DATA_BLOCK "DB_CrossCut_3_HMI"   // DB2078
{ S7_Optimized_Access := 'FALSE' }
VERSION : 0.1
   VAR
      tALM : Struct   // HMI Alarms
         tE : Struct   // Emergency alarms
            xLocON : Bool;   // KE.Local emergency ON {X|X|X|X|O}
            xLocal1 : Bool;   // SB.Local emergency push button 1 {X|X|X|X|O}
            xLocal2 : Bool;   // SB.Local emergency push button 2 {X|X|X|X|O}
            xLocal3 : Bool;   // SB.Local emergency push button 3 {X|X|X|X|O}
            xSpare_4 : Bool;
            xSpare_5 : Bool;
            xSpare_6 : Bool;
            xSpare_7 : Bool;
            xSpare_8 : Bool;
            xSpare_9 : Bool;
            xSpare_10 : Bool;
            xSpare_11 : Bool;
            xSpare_12 : Bool;
            xSpare_13 : Bool;
            xSpare_14 : Bool;
            xSpare_15 : Bool;
            xSpare_16 : Bool;
            xSpare_17 : Bool;
            xSpare_18 : Bool;
            xSpare_19 : Bool;
            xSpare_20 : Bool;
            xSpare_21 : Bool;
            xSpare_22 : Bool;
            xSpare_23 : Bool;
            xSpare_24 : Bool;
            xSpare_25 : Bool;
            xSpare_26 : Bool;
            xSpare_27 : Bool;
            xSpare_28 : Bool;
            xSpare_29 : Bool;
            xSpare_30 : Bool;
            xSpare_31 : Bool;
         END_STRUCT;
         tS : Struct   // Stopping faults
            xAxisNotAvail : Bool;   // AZ.Axis not available {X|X|X|X|O}
            xInpInstallation : Bool;   // L+.Input power supply ON {X|X|X|X|O}
            xAuxPower : Bool;   // L+.Auxiliary power supple set-in {X|X|X|X|O}
            xAreaSafety : Bool;   // KE.Area safety {X|X|X|X|O}
            xOverstroke : Bool;   // KA.Carriage overstroke {X|X|X|X|O}
            xExternInputPower : Bool;   // L+.External input power supply {X|X|X|X|O}
            xCarriageCutOut : Bool;   // QM.Carriage translation overload {X|X|X|X|O}
            xDriveTrip : Bool;   // AZ.Drive trip {X|X|X|X|O}
            xDriveNotEnabled : Bool;   // AZ.Drive not enabled {X|X|X|X|O}
            xAxisNotReady : Bool;   // AZ.Axis not ready {X|X|X|X|O}
            xDriveNotReady : Bool;   // AZ.Drive not ready {X|X|X|X|O}
            xAxisNotSyncro : Bool;   // AZ.Axis not syncronized {X|X|X|X|O}
            xSpare_12 : Bool;
            xSpare_13 : Bool;
            xSpare_14 : Bool;
            xSpare_15 : Bool;
            xSpare_16 : Bool;
            xSpare_17 : Bool;
            xSpare_18 : Bool;
            xSpare_19 : Bool;
            xSpare_20 : Bool;
            xSpare_21 : Bool;
            xSpare_22 : Bool;
            xSpare_23 : Bool;
            xSpare_24 : Bool;
            xSpare_25 : Bool;
            xSpare_26 : Bool;
            xSpare_27 : Bool;
            xSpare_28 : Bool;
            xSpare_29 : Bool;
            xSpare_30 : Bool;
            xSpare_31 : Bool;
         END_STRUCT;
         tF : Struct   // Faults
            xSpare_0 : Bool;
            xSpare_1 : Bool;
            xSpare_2 : Bool;
            xSpare_3 : Bool;
            xSpare_4 : Bool;
            xSpare_5 : Bool;
            xSpare_6 : Bool;
            xSpare_7 : Bool;
            xSpare_8 : Bool;
            xSpare_9 : Bool;
            xSpare_10 : Bool;
            xSpare_11 : Bool;
            xSpare_12 : Bool;
            xSpare_13 : Bool;
            xSpare_14 : Bool;
            xSpare_15 : Bool;
            xSpare_16 : Bool;
            xSpare_17 : Bool;
            xSpare_18 : Bool;
            xSpare_19 : Bool;
            xSpare_20 : Bool;
            xSpare_21 : Bool;
            xSpare_22 : Bool;
            xSpare_23 : Bool;
            xSpare_24 : Bool;
            xSpare_25 : Bool;
            xSpare_26 : Bool;
            xSpare_27 : Bool;
            xSpare_28 : Bool;
            xSpare_29 : Bool;
            xSpare_30 : Bool;
            xSpare_31 : Bool;
         END_STRUCT;
         tW : Struct   // Warnings
            xSpare_0 : Bool;
            xSpare_1 : Bool;
            xSpare_2 : Bool;
            xSpare_3 : Bool;
            xSpare_4 : Bool;
            xSpare_5 : Bool;
            xSpare_6 : Bool;
            xSpare_7 : Bool;
            xSpare_8 : Bool;
            xSpare_9 : Bool;
            xSpare_10 : Bool;
            xSpare_11 : Bool;
            xSpare_12 : Bool;
            xSpare_13 : Bool;
            xSpare_14 : Bool;
            xSpare_15 : Bool;
            xSpare_16 : Bool;
            xSpare_17 : Bool;
            xSpare_18 : Bool;
            xSpare_19 : Bool;
            xSpare_20 : Bool;
            xSpare_21 : Bool;
            xSpare_22 : Bool;
            xSpare_23 : Bool;
            xSpare_24 : Bool;
            xSpare_25 : Bool;
            xSpare_26 : Bool;
            xSpare_27 : Bool;
            xSpare_28 : Bool;
            xSpare_29 : Bool;
            xSpare_30 : Bool;
            xSpare_31 : Bool;
         END_STRUCT;
      END_STRUCT;
      tHMR : Struct   // HMI Read
         xSpare0 : Bool;
         xSpare1 : Bool;
         xSpare2 : Bool;
         xSpare3 : Bool;
         xSpare4 : Bool;
         xSpare5 : Bool;
         xSpare6 : Bool;
         xSpare7 : Bool;
         xSpare8 : Bool;
         xSpare9 : Bool;
         xSpare10 : Bool;
         xSpare11 : Bool;
         xSpare12 : Bool;
         xSpare13 : Bool;
         xManualCommandEnabled : Bool;   // Manual Command enabled {x|x|x|x|O}
         xSpare15 : Bool;
         xSpare16 : Bool;
         xSpare17 : Bool;
         xSpare18 : Bool;
         xSpare19 : Bool;
         xSpare20 : Bool;
         xSpare21 : Bool;
         xSpare22 : Bool;
         xSpare23 : Bool;
         xSpare24 : Bool;
         xSpare25 : Bool;
         xSpare26 : Bool;
         xSpare27 : Bool;
         xSpare28 : Bool;
         xSpare29 : Bool;
         xSpare30 : Bool;
         xSpare31 : Bool;
         xSpare : Array[0..15] of Bool;
         iSpare0 : Int;
         iSpare1 : Int;
         iSpare2 : Int;
         iSpare3 : Int;
         iSpare4 : Int;
         iSpare5 : Int;
         iSpare6 : Int;
         iSpare7 : Int;
         iSpare8 : Int;
         iSpare9 : Int;
         iSpare10 : Int;
         iSpare11 : Int;
         iSpare12 : Int;
         iSpare13 : Int;
         iSpare14 : Int;
         iSpare15 : Int;
         iSpare16 : Int;
         dDistanceSnaproll_cmm : DInt;   // Distance from snaproll [mm/100] {mm/100|mm|x|x|M}
         dStatus : DInt;   // XCut actual status (1=Idle 3=Running 7=Faulted) {X|X|X|X|O}
         dXCutActualStatus : DInt;   // XCut actual status (1=Disabled 3=Enabled) {X|X|X|X|O}
         dXCutStatusRequest : DInt;   // XCut status request (1=Disabled 3=Enabled) {X|X|X|X|O}
         dDistanceFromCenterLine_cmm : DInt;   // Distance from center line [mm/100] {mm/100|mm|X|X|O}
         dAngleValue_uDegree : DInt;   // Angle value [°/1000000] {°/1000000|°|X|X|O}
         dActualCutPosRequest : DInt;   // Actual cut position request (1=By operator 2=On gross ribbon 3=On net ribbon 4=On YCut position) {X|X|X|X|O}
         dCarriagePosition_cmm : DInt;   // Actual carriage position [mm/100]
         dSpare8 : DInt;
         dSpare9 : DInt;
         dSpare10 : DInt;
         dSpare11 : DInt;
         dSpare12 : DInt;
         dSpare13 : DInt;
         dSpare14 : DInt;
         dSpare15 : DInt;
         rHeadUsage_km : Real;   // Head usage [Km] {Km|Km|X|X|O}
         rSpare1 : Real;
         rSpare2 : Real;
         rSpare3 : Real;
         rSpare4 : Real;
         rSpare5 : Real;
         rSpare6 : Real;
         rSpare7 : Real;
         rSpare8 : Real;
         tManCmd : Struct
            xManJogFwdFdbk : Bool;   // Manual jog forward feedback {X|X|X|X|O}
            xManJogBckFdbk : Bool;   // Manual jog backward feedback {X|X|X|X|O}
            xManCarriageDownFdbk : Bool;   // Manual carriage down feedback {X|X|X|X|O}
            xManFireONFdbk : Bool;   // Manual fire ON feedback {X|X|X|X|O}
            xManOilONFdbk : Bool;   // Manual oil ON feedback {X|X|X|X|O}
            xSpare5 : Bool;
            xSpare6 : Bool;
            xSpare7 : Bool;
            xSpare8 : Bool;
            xSpare9 : Bool;
            xSpare10 : Bool;
            xSpare11 : Bool;
            xSpare12 : Bool;
            xSpare13 : Bool;
            xSpare14 : Bool;
            xSpare15 : Bool;
            xSpare : Array[0..15] of Bool;
         END_STRUCT;
      END_STRUCT;
      tHMW : Struct   // HMI Write
         xCutBreakEnabled : Bool;   // Cut on glass break enabled {X|X|X|X|O}
         xIncAngleValue : Bool;   // Increment angle value {X|X|X|X|O}
         xDecAngleValue : Bool;   // Decrement angle value {X|X|X|X|O}
         xCalibDistRequest : Bool;   // Calibration distance request {X|X|X|X|O}
         xCalibDiagRequest : Bool;   // Calibration diagonal request {X|X|X|X|O}
         xCutOperator : Bool;   // Cutting position by operator request {X|X|X|X|O}
         xCutGross : Bool;   // Cutting position by gross width position {X|X|X|X|O}
         xCutNet : Bool;   // Cutting position by net width position {X|X|X|X|O}
         xCutYCut : Bool;   // Cutting position by YCut position {X|X|X|X|O}
         xSpare9 : Bool;
         xSpare10 : Bool;
         xSpare11 : Bool;
         xSpare12 : Bool;
         xResetHeadUsage : Bool;   // Reset the head usage {X|X|X|X|O}
         xEnableManualCommand : Bool;   // Enable Disable Manual command {x|x|x|x|O}
         xUpdateDistanceSnaproll : Bool;   // Update distance from snaproll {x|x|x|x|M}
         xUpdateDistCenterLine : Bool;   // Update distance from center line {X|X|X|X|M}
         xUpdateAngleValue : Bool;   // Update angle value {X|X|X|X|M}
         xSpare18 : Bool;
         xSpare19 : Bool;
         xSpare20 : Bool;
         xSpare21 : Bool;
         xSpare22 : Bool;
         xSpare23 : Bool;
         xSpare24 : Bool;
         xSpare25 : Bool;
         xSpare26 : Bool;
         xSpare27 : Bool;
         xSpare28 : Bool;
         xSpare29 : Bool;
         xSpare30 : Bool;
         xSpare31 : Bool;
         xSpare : Array[0..15] of Bool;
         iSpare0 : Int;
         iSpare1 : Int;
         iSpare2 : Int;
         iSpare3 : Int;
         iSpare4 : Int;
         iSpare5 : Int;
         iSpare6 : Int;
         iSpare7 : Int;
         iSpare8 : Int;
         iSpare9 : Int;
         iSpare10 : Int;
         iSpare11 : Int;
         iSpare12 : Int;
         iSpare13 : Int;
         iSpare14 : Int;
         iSpare15 : Int;
         iSpare16 : Int;
         dDistanceSnaproll_cmm : DInt;   // Distance from snaproll [mm/100] {mm/100|mm|1|70000|M}
         dDistanceFromCenterLine_cmm : DInt;   // Distance from center line [mm/100] {mm/100|mm|-3000|0|M}
         dAngleValue_uDegree : DInt;   // Bridge angle value [°/1000000] {°/1000000|°|7|9|M}
         dOperStartCutPos_cmm : DInt;   // Operator start cut position [mm/100] {mm/100|mm|-3000|0|O}
         dOperEndCutPos_cmm : DInt;   // Operator end cut position [mm/100] {mm/100|mm|0|3000|O}
         dDescReactTime_ms : DInt;   // Carriage descent reaction time [ms] {ms|s|0|1|M}
         dRaiseReactTime_ms : DInt;   // Carriage raise reaction time [ms] {ms|s|0|1|M}
         dFireONReactTime_ms : DInt;   // Fire ON reaction time [ms] {ms|s|0|1|M}
         dFireOFFReactTime_ms : DInt;   // Fire OFF reaction time [ms] {ms|s|0|1|M}
         dOilONDelay_ms : DInt;   // Oil ON delay [ms] {ms|s|-1|1|O}
         dOilOFFDelay_ms : DInt;   // Oil OFF delay [ms] {ms|s|-1|1|O}
         dCutStartOffsetDelay_cmm : DInt;   // Start cut offset delay [mm/100] {mm/100|mm|-500|500|O}
         dCutEndOffsetDelay_cmm : DInt;   // End cut offset delay [mm/100] {mm/100|mm|-500|500|O}
         dDistTeoLength_cmm : DInt;   // Calibration distance.Theorical length [mm/100] {mm/100|mm|0|7000|O}
         dDistRealLength_cmm : DInt;   // Calibration distance.Real length [mm/100] {mm/100|mm|0|7000|O}
         dDiagRealLength_cmm : DInt;   // Calibration diagonal.Real length [mm/100] {mm/100|mm|0|7000|O}
         dDiagRealWidth_cmm : DInt;   // Calibration diagonal.Real width [mm/100] {mm/100|mm|0|4000|O}
         dDiagGlassFlow_cmm : DInt;   // Calibration diagonal.Real length diagonal glass flow [mm/100] {mm/100|mm|0|10000|O}
         dDiagGlassOppFlow_cmm : DInt;   // Calibration diagonal.Real length diagonal opposite glass flow [mm/100] {mm/100|mm|0|10000|O}
         dCuttingPressure_mN : DInt;   // Cutting pressure [N/1000] {N/1000|N|9|180|O}
         dPosOffset_cmm : DInt;   // Calibration offset distance from snaproll [mm/100] {mm/100|mm|-50|50|O}
         dCutPriority : DInt;   // Cut priority number {X|X|0|5|O}
         dSpare22 : DInt;
         rSpare6 : Real;
         rSpare7 : Real;
         rSpare8 : Real;
         tManCmd : Struct
            xMan_JogForward : Bool;   // Manual mode - Jog forward {X|X|X|X|M}
            xMan_JobBackward : Bool;   // Manual mode - Jog backward {X|X|X|X|M}
            xMan_CarriageDown : Bool;   // Manual mode - Carriage down {X|X|X|X|M}
            xMan_FireOn : Bool;   // Manual mode - Fire ON {X|X|X|X|M}
            xMan_OilOn : Bool;   // Manual mode - Oil ON {X|X|X|X|M}
            xSpare5 : Bool;
            xSpare6 : Bool;
            xSpare7 : Bool;
            xSpare8 : Bool;
            xSpare9 : Bool;
            xSpare10 : Bool;
            xSpare11 : Bool;
            xSpare12 : Bool;
            xSpare13 : Bool;
            xSpare14 : Bool;
            xSpare15 : Bool;
            xSpare16 : Bool;
            xSpare17 : Bool;
            xSpare18 : Bool;
            xSpare19 : Bool;
            xSpare20 : Bool;
            xSpare21 : Bool;
            xSpare22 : Bool;
            xSpare23 : Bool;
            xSpare24 : Bool;
            xSpare25 : Bool;
            xSpare26 : Bool;
            xSpare27 : Bool;
            xSpare28 : Bool;
            xSpare29 : Bool;
            xSpare30 : Bool;
            xSpare31 : Bool;
         END_STRUCT;
      END_STRUCT;
   END_VAR
BEGIN
END_DATA_BLOCK

DATA_BLOCK "DB_Marker_HMI"   // DB2081
{ S7_Optimized_Access := 'FALSE' }
VERSION : 0.1
   VAR
      tALM : Struct   // HMI Alarms
         tE : Struct   // Stopping faults
            xSpare_0 : Bool;
            xSpare_1 : Bool;
            xSpare_2 : Bool;
            xSpare_3 : Bool;
            xSpare_4 : Bool;
            xSpare_5 : Bool;
            xSpare_6 : Bool;
            xSpare_7 : Bool;
            xSpare_8 : Bool;
            xSpare_9 : Bool;
            xSpare_10 : Bool;
            xSpare_11 : Bool;
            xSpare_12 : Bool;
            xSpare_13 : Bool;
            xSpare_14 : Bool;
            xSpare_15 : Bool;
            xSpare_16 : Bool;
            xSpare_17 : Bool;
            xSpare_18 : Bool;
            xSpare_19 : Bool;
            xSpare_20 : Bool;
            xSpare_21 : Bool;
            xSpare_22 : Bool;
            xSpare_23 : Bool;
            xSpare_24 : Bool;
            xSpare_25 : Bool;
            xSpare_26 : Bool;
            xSpare_27 : Bool;
            xSpare_28 : Bool;
            xSpare_29 : Bool;
            xSpare_30 : Bool;
            xSpare_31 : Bool;
         END_STRUCT;
         tS : Struct   // Stopping faults
            xTOutSendData : Bool;   // Timeout send data to bridge
            xSpare_1 : Bool;
            xSpare_2 : Bool;
            xSpare_3 : Bool;
            xSpare_4 : Bool;
            xSpare_5 : Bool;
            xSpare_6 : Bool;
            xSpare_7 : Bool;
            xSpare_8 : Bool;
            xSpare_9 : Bool;
            xSpare_10 : Bool;
            xSpare_11 : Bool;
            xSpare_12 : Bool;
            xSpare_13 : Bool;
            xSpare_14 : Bool;
            xSpare_15 : Bool;
            xSpare_16 : Bool;
            xSpare_17 : Bool;
            xSpare_18 : Bool;
            xSpare_19 : Bool;
            xSpare_20 : Bool;
            xSpare_21 : Bool;
            xSpare_22 : Bool;
            xSpare_23 : Bool;
            xSpare_24 : Bool;
            xSpare_25 : Bool;
            xSpare_26 : Bool;
            xSpare_27 : Bool;
            xSpare_28 : Bool;
            xSpare_29 : Bool;
            xSpare_30 : Bool;
            xSpare_31 : Bool;
         END_STRUCT;
         tF : Struct   // Faults
            xSpare_0 : Bool;
            xSpare_1 : Bool;
            xSpare_2 : Bool;
            xSpare_3 : Bool;
            xSpare_4 : Bool;
            xSpare_5 : Bool;
            xSpare_6 : Bool;
            xSpare_7 : Bool;
            xSpare_8 : Bool;
            xSpare_9 : Bool;
            xSpare_10 : Bool;
            xSpare_11 : Bool;
            xSpare_12 : Bool;
            xSpare_13 : Bool;
            xSpare_14 : Bool;
            xSpare_15 : Bool;
            xSpare_16 : Bool;
            xSpare_17 : Bool;
            xSpare_18 : Bool;
            xSpare_19 : Bool;
            xSpare_20 : Bool;
            xSpare_21 : Bool;
            xSpare_22 : Bool;
            xSpare_23 : Bool;
            xSpare_24 : Bool;
            xSpare_25 : Bool;
            xSpare_26 : Bool;
            xSpare_27 : Bool;
            xSpare_28 : Bool;
            xSpare_29 : Bool;
            xSpare_30 : Bool;
            xSpare_31 : Bool;
         END_STRUCT;
         tW : Struct   // Warnings
            xSpare_0 : Bool;
            xSpare_1 : Bool;
            xSpare_2 : Bool;
            xSpare_3 : Bool;
            xSpare_4 : Bool;
            xSpare_5 : Bool;
            xSpare_6 : Bool;
            xSpare_7 : Bool;
            xSpare_8 : Bool;
            xSpare_9 : Bool;
            xSpare_10 : Bool;
            xSpare_11 : Bool;
            xSpare_12 : Bool;
            xSpare_13 : Bool;
            xSpare_14 : Bool;
            xSpare_15 : Bool;
            xSpare_16 : Bool;
            xSpare_17 : Bool;
            xSpare_18 : Bool;
            xSpare_19 : Bool;
            xSpare_20 : Bool;
            xSpare_21 : Bool;
            xSpare_22 : Bool;
            xSpare_23 : Bool;
            xSpare_24 : Bool;
            xSpare_25 : Bool;
            xSpare_26 : Bool;
            xSpare_27 : Bool;
            xSpare_28 : Bool;
            xSpare_29 : Bool;
            xSpare_30 : Bool;
            xSpare_31 : Bool;
         END_STRUCT;
      END_STRUCT;
      tHMR : Struct   // HMI Read
         xSpare0 : Bool;
         xSpare1 : Bool;
         xSpare2 : Bool;
         xSpare3 : Bool;
         xSpare4 : Bool;
         xSpare5 : Bool;
         xSpare6 : Bool;
         xSpare7 : Bool;
         xSpare8 : Bool;
         xSpare9 : Bool;
         xSpare10 : Bool;
         xSpare11 : Bool;
         xSpare12 : Bool;
         xSpare13 : Bool;
         xSpare14 : Bool;
         xSpare15 : Bool;
         xSpare16 : Bool;
         xSpare17 : Bool;
         xSpare18 : Bool;
         xSpare19 : Bool;
         xSpare20 : Bool;
         xSpare21 : Bool;
         xSpare22 : Bool;
         xSpare23 : Bool;
         xSpare24 : Bool;
         xSpare25 : Bool;
         xSpare26 : Bool;
         xSpare27 : Bool;
         xSpare28 : Bool;
         xSpare29 : Bool;
         xSpare30 : Bool;
         xSpare31 : Bool;
         xSpare : Array[0..15] of Bool;
         iSpare0 : Int;
         iSpare1 : Int;
         iSpare2 : Int;
         iSpare3 : Int;
         iSpare4 : Int;
         iSpare5 : Int;
         iSpare6 : Int;
         iSpare7 : Int;
         iSpare8 : Int;
         iSpare9 : Int;
         iSpare10 : Int;
         iSpare11 : Int;
         iSpare12 : Int;
         iSpare13 : Int;
         iSpare14 : Int;
         iSpare15 : Int;
         iSpare16 : Int;
         dSpare0 : DInt;
         dSpare1 : DInt;
         dSpare2 : DInt;
         dSpare3 : DInt;
         dSpare4 : DInt;
         dSpare5 : DInt;
         dSpare6 : DInt;
         dSpare7 : DInt;
         dSpare8 : DInt;
         dSpare9 : DInt;
         dSpare10 : DInt;
         dSpare11 : DInt;
         dSpare12 : DInt;
         dSpare13 : DInt;
         dSpare14 : DInt;
         dSpare15 : DInt;
         rSpare0 : Real;
         rSpare1 : Real;
         rSpare2 : Real;
         rSpare3 : Real;
         rSpare4 : Real;
         rSpare5 : Real;
         rSpare6 : Real;
         rSpare7 : Real;
         rSpare8 : Real;
         tManCmd : Struct
            xSpare0 : Bool;
            xSpare1 : Bool;
            xSpare2 : Bool;
            xSpare3 : Bool;
            xSpare4 : Bool;
            xSpare5 : Bool;
            xSpare6 : Bool;
            xSpare7 : Bool;
            xSpare8 : Bool;
            xSpare9 : Bool;
            xSpare10 : Bool;
            xSpare11 : Bool;
            xSpare12 : Bool;
            xSpare13 : Bool;
            xSpare14 : Bool;
            xSpare15 : Bool;
            xSpare : Array[0..15] of Bool;
         END_STRUCT;
      END_STRUCT;
      tHMW : Struct   // HMI Write
         xSpare0 : Bool;
         xSpare1 : Bool;
         xSpare2 : Bool;
         xSpare3 : Bool;
         xSpare4 : Bool;
         xSpare5 : Bool;
         xSpare6 : Bool;
         xSpare7 : Bool;
         xSpare8 : Bool;
         xSpare9 : Bool;
         xSpare10 : Bool;
         xSpare11 : Bool;
         xSpare12 : Bool;
         xSpare13 : Bool;
         xSpare14 : Bool;
         xSpare15 : Bool;
         xSpare16 : Bool;
         xSpare17 : Bool;
         xSpare18 : Bool;
         xSpare19 : Bool;
         xSpare20 : Bool;
         xSpare21 : Bool;
         xSpare22 : Bool;
         xSpare23 : Bool;
         xSpare24 : Bool;
         xSpare25 : Bool;
         xSpare26 : Bool;
         xSpare27 : Bool;
         xSpare28 : Bool;
         xSpare29 : Bool;
         xSpare30 : Bool;
         xSpare31 : Bool;
         xSpare : Array[0..15] of Bool;
         iSpare0 : Int;
         iSpare1 : Int;
         iSpare2 : Int;
         iSpare3 : Int;
         iSpare4 : Int;
         iSpare5 : Int;
         iSpare6 : Int;
         iSpare7 : Int;
         iSpare8 : Int;
         iSpare9 : Int;
         iSpare10 : Int;
         iSpare11 : Int;
         iSpare12 : Int;
         iSpare13 : Int;
         iSpare14 : Int;
         iSpare15 : Int;
         iSpare16 : Int;
         dSpare0 : DInt;
         dSpare1 : DInt;
         dSpare2 : DInt;
         dSpare3 : DInt;
         dSpare4 : DInt;
         dSpare5 : DInt;
         dSpare6 : DInt;
         dSpare7 : DInt;
         dSpare8 : DInt;
         dSpare9 : DInt;
         dSpare10 : DInt;
         dSpare11 : DInt;
         dSpare12 : DInt;
         dSpare13 : DInt;
         dSpare14 : DInt;
         dSpare15 : DInt;
         dSpare16 : DInt;
         rSpare0 : Real;
         rSpare1 : Real;
         rSpare2 : Real;
         rSpare3 : Real;
         rSpare4 : Real;
         rSpare5 : Real;
         rSpare6 : Real;
         rSpare7 : Real;
         rSpare8 : Real;
         tManCmd : Struct
            xSpare0 : Bool;
            xSpare1 : Bool;
            xSpare2 : Bool;
            xSpare3 : Bool;
            xSpare4 : Bool;
            xSpare5 : Bool;
            xSpare6 : Bool;
            xSpare7 : Bool;
            xSpare8 : Bool;
            xSpare9 : Bool;
            xSpare10 : Bool;
            xSpare11 : Bool;
            xSpare12 : Bool;
            xSpare13 : Bool;
            xSpare14 : Bool;
            xSpare15 : Bool;
            xSpare16 : Bool;
            xSpare17 : Bool;
            xSpare18 : Bool;
            xSpare19 : Bool;
            xSpare20 : Bool;
            xSpare21 : Bool;
            xSpare22 : Bool;
            xSpare23 : Bool;
            xSpare24 : Bool;
            xSpare25 : Bool;
            xSpare26 : Bool;
            xSpare27 : Bool;
            xSpare28 : Bool;
            xSpare29 : Bool;
            xSpare30 : Bool;
            xSpare31 : Bool;
         END_STRUCT;
      END_STRUCT;
   END_VAR
BEGIN
END_DATA_BLOCK

DATA_BLOCK "DB_SnapRoll_221_HMI"   // DB2095
{ S7_Optimized_Access := 'FALSE' }
VERSION : 0.1
   VAR
      tALM : Struct   // HMI Alarms
         tE : Struct   // Stopping faults
            xSpare_0 : Bool;
            xSpare_1 : Bool;
            xSpare_2 : Bool;
            xSpare_3 : Bool;
            xSpare_4 : Bool;
            xSpare_5 : Bool;
            xSpare_6 : Bool;
            xSpare_7 : Bool;
            xSpare_8 : Bool;
            xSpare_9 : Bool;
            xSpare_10 : Bool;
            xSpare_11 : Bool;
            xSpare_12 : Bool;
            xSpare_13 : Bool;
            xSpare_14 : Bool;
            xSpare_15 : Bool;
            xSpare_16 : Bool;
            xSpare_17 : Bool;
            xSpare_18 : Bool;
            xSpare_19 : Bool;
            xSpare_20 : Bool;
            xSpare_21 : Bool;
            xSpare_22 : Bool;
            xSpare_23 : Bool;
            xSpare_24 : Bool;
            xSpare_25 : Bool;
            xSpare_26 : Bool;
            xSpare_27 : Bool;
            xSpare_28 : Bool;
            xSpare_29 : Bool;
            xSpare_30 : Bool;
            xSpare_31 : Bool;
         END_STRUCT;
         tS : Struct   // Stopping faults
            xSpare_0 : Bool;
            xSpare_1 : Bool;
            xSpare_2 : Bool;
            xSpare_3 : Bool;
            xSpare_4 : Bool;
            xSpare_5 : Bool;
            xSpare_6 : Bool;
            xSpare_7 : Bool;
            xSpare_8 : Bool;
            xSpare_9 : Bool;
            xSpare_10 : Bool;
            xSpare_11 : Bool;
            xSpare_12 : Bool;
            xSpare_13 : Bool;
            xSpare_14 : Bool;
            xSpare_15 : Bool;
            xSpare_16 : Bool;
            xSpare_17 : Bool;
            xSpare_18 : Bool;
            xSpare_19 : Bool;
            xSpare_20 : Bool;
            xSpare_21 : Bool;
            xSpare_22 : Bool;
            xSpare_23 : Bool;
            xSpare_24 : Bool;
            xSpare_25 : Bool;
            xSpare_26 : Bool;
            xSpare_27 : Bool;
            xSpare_28 : Bool;
            xSpare_29 : Bool;
            xSpare_30 : Bool;
            xSpare_31 : Bool;
         END_STRUCT;
         tF : Struct   // Faults
            xSpare_0 : Bool;
            xSpare_1 : Bool;
            xSpare_2 : Bool;
            xSpare_3 : Bool;
            xSpare_4 : Bool;
            xSpare_5 : Bool;
            xSpare_6 : Bool;
            xSpare_7 : Bool;
            xSpare_8 : Bool;
            xSpare_9 : Bool;
            xSpare_10 : Bool;
            xSpare_11 : Bool;
            xSpare_12 : Bool;
            xSpare_13 : Bool;
            xSpare_14 : Bool;
            xSpare_15 : Bool;
            xSpare_16 : Bool;
            xSpare_17 : Bool;
            xSpare_18 : Bool;
            xSpare_19 : Bool;
            xSpare_20 : Bool;
            xSpare_21 : Bool;
            xSpare_22 : Bool;
            xSpare_23 : Bool;
            xSpare_24 : Bool;
            xSpare_25 : Bool;
            xSpare_26 : Bool;
            xSpare_27 : Bool;
            xSpare_28 : Bool;
            xSpare_29 : Bool;
            xSpare_30 : Bool;
            xSpare_31 : Bool;
         END_STRUCT;
         tW : Struct   // Warnings
            xSpare_0 : Bool;
            xSpare_1 : Bool;
            xSpare_2 : Bool;
            xSpare_3 : Bool;
            xSpare_4 : Bool;
            xSpare_5 : Bool;
            xSpare_6 : Bool;
            xSpare_7 : Bool;
            xSpare_8 : Bool;
            xSpare_9 : Bool;
            xSpare_10 : Bool;
            xSpare_11 : Bool;
            xSpare_12 : Bool;
            xSpare_13 : Bool;
            xSpare_14 : Bool;
            xSpare_15 : Bool;
            xSpare_16 : Bool;
            xSpare_17 : Bool;
            xSpare_18 : Bool;
            xSpare_19 : Bool;
            xSpare_20 : Bool;
            xSpare_21 : Bool;
            xSpare_22 : Bool;
            xSpare_23 : Bool;
            xSpare_24 : Bool;
            xSpare_25 : Bool;
            xSpare_26 : Bool;
            xSpare_27 : Bool;
            xSpare_28 : Bool;
            xSpare_29 : Bool;
            xSpare_30 : Bool;
            xSpare_31 : Bool;
         END_STRUCT;
      END_STRUCT;
      tHMR : Struct   // HMI Read
         xSpare0 : Bool;
         xSpare1 : Bool;
         xSpare2 : Bool;
         xSpare3 : Bool;
         xSpare4 : Bool;
         xSpare5 : Bool;
         xSpare6 : Bool;
         xSpare7 : Bool;
         xSpare8 : Bool;
         xSpare9 : Bool;
         xSpare10 : Bool;
         xSpare11 : Bool;
         xSpare12 : Bool;
         xSpare13 : Bool;
         xManualCommandEnabled : Bool;   // Manual Command enabled {x|x|x|x|O}
         xSpare15 : Bool;
         xSpare16 : Bool;
         xSpare17 : Bool;
         xSpare18 : Bool;
         xSpare19 : Bool;
         xSpare20 : Bool;
         xSpare21 : Bool;
         xSpare22 : Bool;
         xSpare23 : Bool;
         xSpare24 : Bool;
         xSpare25 : Bool;
         xSpare26 : Bool;
         xSpare27 : Bool;
         xSpare28 : Bool;
         xSpare29 : Bool;
         xSpare30 : Bool;
         xSpare31 : Bool;
         xSpare : Array[0..15] of Bool;
         iSpare0 : Int;
         iSpare1 : Int;
         iSpare2 : Int;
         iSpare3 : Int;
         iSpare4 : Int;
         iSpare5 : Int;
         iSpare6 : Int;
         iSpare7 : Int;
         iSpare8 : Int;
         iSpare9 : Int;
         iSpare10 : Int;
         iSpare11 : Int;
         iSpare12 : Int;
         iSpare13 : Int;
         iSpare14 : Int;
         iSpare15 : Int;
         iSpare16 : Int;
         dSpare0 : DInt;
         dStatus : DInt;   // Status (1=Idle 3=Up 7=Fault) {x|x|x|x|O}
         dSpare2 : DInt;
         dSpare3 : DInt;
         dSpare4 : DInt;
         dSpare5 : DInt;
         dSpare6 : DInt;
         dSpare7 : DInt;
         dSpare8 : DInt;
         dSpare9 : DInt;
         dSpare10 : DInt;
         dSpare11 : DInt;
         dSpare12 : DInt;
         dSpare13 : DInt;
         dSpare14 : DInt;
         dSpare15 : DInt;
         rSpare0 : Real;
         rSpare1 : Real;
         rSpare2 : Real;
         rSpare3 : Real;
         rSpare4 : Real;
         rSpare5 : Real;
         rSpare6 : Real;
         rSpare7 : Real;
         rSpare8 : Real;
         tManCmd : Struct
            xUp : Bool;   // Snap roll up feedback {x|x|x|x|O}
            xContrastActivation : Bool;   // Contrast activation feedback {x|x|x|x|O}
            xSpare2 : Bool;
            xSpare3 : Bool;
            xSpare4 : Bool;
            xSpare5 : Bool;
            xSpare6 : Bool;
            xSpare7 : Bool;
            xSpare8 : Bool;
            xSpare9 : Bool;
            xSpare10 : Bool;
            xSpare11 : Bool;
            xSpare12 : Bool;
            xSpare13 : Bool;
            xSpare14 : Bool;
            xSpare15 : Bool;
            xSpare : Array[0..15] of Bool;
         END_STRUCT;
      END_STRUCT;
      tHMW : Struct   // HMI Write
         xSpare0 : Bool;
         xSpare1 : Bool;
         xSpare2 : Bool;
         xSpare3 : Bool;
         xSpare4 : Bool;
         xSpare5 : Bool;
         xSpare6 : Bool;
         xSpare7 : Bool;
         xSpare8 : Bool;
         xSpare9 : Bool;
         xSpare10 : Bool;
         xSpare11 : Bool;
         xSpare12 : Bool;
         xSpare13 : Bool;
         xEnableManualCommand : Bool;   // Enable Disable Manual command {x|x|x|x|O}
         xSpare15 : Bool;
         xSpare16 : Bool;
         xSpare17 : Bool;
         xSpare18 : Bool;
         xSpare19 : Bool;
         xSpare20 : Bool;
         xSpare21 : Bool;
         xSpare22 : Bool;
         xSpare23 : Bool;
         xSpare24 : Bool;
         xSpare25 : Bool;
         xSpare26 : Bool;
         xSpare27 : Bool;
         xSpare28 : Bool;
         xSpare29 : Bool;
         xSpare30 : Bool;
         xSpare31 : Bool;
         xSpare : Array[0..15] of Bool;
         iSpare0 : Int;
         iSpare1 : Int;
         iSpare2 : Int;
         iSpare3 : Int;
         iSpare4 : Int;
         iSpare5 : Int;
         iSpare6 : Int;
         iSpare7 : Int;
         iSpare8 : Int;
         iSpare9 : Int;
         iSpare10 : Int;
         iSpare11 : Int;
         iSpare12 : Int;
         iSpare13 : Int;
         iSpare14 : Int;
         iSpare15 : Int;
         iSpare16 : Int;
         dOffsetSnap_cmm : DInt;   // Offset rise snap (- Anticipate + Delay) [mm/100] {mm/100|mm|-300|300|O}
         dMaxPlateLenghtEnableContrast_cmm : DInt;   // Maximum plate lenght for contrast enabling [mm/100] {mm/100|mm|1|7000|O}
         dTimeUp_ms : DInt;   // Time snap in up position [ms] {ms|s|0|1|O}
         dReactTime_ms : DInt;   // Snap reaction time [ms] {ms|s|0|1|O}
         dSpare4 : DInt;
         dSpare5 : DInt;
         dSpare6 : DInt;
         dSpare7 : DInt;
         dSpare8 : DInt;
         dSpare9 : DInt;
         dSpare10 : DInt;
         dSpare11 : DInt;
         dSpare12 : DInt;
         dSpare13 : DInt;
         dSpare14 : DInt;
         dSpare15 : DInt;
         dSpare16 : DInt;
         rSpare0 : Real;
         rSpare1 : Real;
         rSpare2 : Real;
         rSpare3 : Real;
         rSpare4 : Real;
         rSpare5 : Real;
         rSpare6 : Real;
         rSpare7 : Real;
         rSpare8 : Real;
         tManCmd : Struct
            xUp : Bool;   // Snap roll up {x|x|x|x|O}
            xContrastActivation : Bool;   // Contrast activation {x|x|x|x|O}
            xSpare2 : Bool;
            xSpare3 : Bool;
            xSpare4 : Bool;
            xSpare5 : Bool;
            xSpare6 : Bool;
            xSpare7 : Bool;
            xSpare8 : Bool;
            xSpare9 : Bool;
            xSpare10 : Bool;
            xSpare11 : Bool;
            xSpare12 : Bool;
            xSpare13 : Bool;
            xSpare14 : Bool;
            xSpare15 : Bool;
            xSpare16 : Bool;
            xSpare17 : Bool;
            xSpare18 : Bool;
            xSpare19 : Bool;
            xSpare20 : Bool;
            xSpare21 : Bool;
            xSpare22 : Bool;
            xSpare23 : Bool;
            xSpare24 : Bool;
            xSpare25 : Bool;
            xSpare26 : Bool;
            xSpare27 : Bool;
            xSpare28 : Bool;
            xSpare29 : Bool;
            xSpare30 : Bool;
            xSpare31 : Bool;
         END_STRUCT;
      END_STRUCT;
   END_VAR
BEGIN
END_DATA_BLOCK

DATA_BLOCK "DB_BPS_A_HMI"   // DB2110
{ S7_Optimized_Access := 'FALSE' }
VERSION : 0.1
   VAR
      tALM : Struct   // HMI Alarms
         tE : Struct   // Stopping faults
            xSpare_0 : Bool;
            xSpare_1 : Bool;
            xSpare_2 : Bool;
            xSpare_3 : Bool;
            xSpare_4 : Bool;
            xSpare_5 : Bool;
            xSpare_6 : Bool;
            xSpare_7 : Bool;
            xSpare_8 : Bool;
            xSpare_9 : Bool;
            xSpare_10 : Bool;
            xSpare_11 : Bool;
            xSpare_12 : Bool;
            xSpare_13 : Bool;
            xSpare_14 : Bool;
            xSpare_15 : Bool;
            xSpare_16 : Bool;
            xSpare_17 : Bool;
            xSpare_18 : Bool;
            xSpare_19 : Bool;
            xSpare_20 : Bool;
            xSpare_21 : Bool;
            xSpare_22 : Bool;
            xSpare_23 : Bool;
            xSpare_24 : Bool;
            xSpare_25 : Bool;
            xSpare_26 : Bool;
            xSpare_27 : Bool;
            xSpare_28 : Bool;
            xSpare_29 : Bool;
            xSpare_30 : Bool;
            xSpare_31 : Bool;
         END_STRUCT;
         tS : Struct   // Stopping faults
            xTimeOutSendBPSData : Bool;   // Time out send BPS data
            xSpare_1 : Bool;
            xSpare_2 : Bool;
            xSpare_3 : Bool;
            xSpare_4 : Bool;
            xSpare_5 : Bool;
            xSpare_6 : Bool;
            xSpare_7 : Bool;
            xSpare_8 : Bool;
            xSpare_9 : Bool;
            xSpare_10 : Bool;
            xSpare_11 : Bool;
            xSpare_12 : Bool;
            xSpare_13 : Bool;
            xSpare_14 : Bool;
            xSpare_15 : Bool;
            xSpare_16 : Bool;
            xSpare_17 : Bool;
            xSpare_18 : Bool;
            xSpare_19 : Bool;
            xSpare_20 : Bool;
            xSpare_21 : Bool;
            xSpare_22 : Bool;
            xSpare_23 : Bool;
            xSpare_24 : Bool;
            xSpare_25 : Bool;
            xSpare_26 : Bool;
            xSpare_27 : Bool;
            xSpare_28 : Bool;
            xSpare_29 : Bool;
            xSpare_30 : Bool;
            xSpare_31 : Bool;
         END_STRUCT;
         tF : Struct   // Faults
            xSpare_0 : Bool;
            xSpare_1 : Bool;
            xSpare_2 : Bool;
            xSpare_3 : Bool;
            xSpare_4 : Bool;
            xSpare_5 : Bool;
            xSpare_6 : Bool;
            xSpare_7 : Bool;
            xSpare_8 : Bool;
            xSpare_9 : Bool;
            xSpare_10 : Bool;
            xSpare_11 : Bool;
            xSpare_12 : Bool;
            xSpare_13 : Bool;
            xSpare_14 : Bool;
            xSpare_15 : Bool;
            xSpare_16 : Bool;
            xSpare_17 : Bool;
            xSpare_18 : Bool;
            xSpare_19 : Bool;
            xSpare_20 : Bool;
            xSpare_21 : Bool;
            xSpare_22 : Bool;
            xSpare_23 : Bool;
            xSpare_24 : Bool;
            xSpare_25 : Bool;
            xSpare_26 : Bool;
            xSpare_27 : Bool;
            xSpare_28 : Bool;
            xSpare_29 : Bool;
            xSpare_30 : Bool;
            xSpare_31 : Bool;
         END_STRUCT;
         tW : Struct   // Warnings
            xSpare_0 : Bool;
            xSpare_1 : Bool;
            xSpare_2 : Bool;
            xSpare_3 : Bool;
            xSpare_4 : Bool;
            xSpare_5 : Bool;
            xSpare_6 : Bool;
            xSpare_7 : Bool;
            xSpare_8 : Bool;
            xSpare_9 : Bool;
            xSpare_10 : Bool;
            xSpare_11 : Bool;
            xSpare_12 : Bool;
            xSpare_13 : Bool;
            xSpare_14 : Bool;
            xSpare_15 : Bool;
            xSpare_16 : Bool;
            xSpare_17 : Bool;
            xSpare_18 : Bool;
            xSpare_19 : Bool;
            xSpare_20 : Bool;
            xSpare_21 : Bool;
            xSpare_22 : Bool;
            xSpare_23 : Bool;
            xSpare_24 : Bool;
            xSpare_25 : Bool;
            xSpare_26 : Bool;
            xSpare_27 : Bool;
            xSpare_28 : Bool;
            xSpare_29 : Bool;
            xSpare_30 : Bool;
            xSpare_31 : Bool;
         END_STRUCT;
      END_STRUCT;
      tHMR : Struct   // HMI Read
         xSpare0 : Bool;
         xSpare1 : Bool;
         xSpare2 : Bool;
         xSpare3 : Bool;
         xSpare4 : Bool;
         xSpare5 : Bool;
         xSpare6 : Bool;
         xSpare7 : Bool;
         xSpare8 : Bool;
         xSpare9 : Bool;
         xSpare10 : Bool;
         xSpare11 : Bool;
         xSpare12 : Bool;
         xSpare13 : Bool;
         xSpare14 : Bool;
         xSpare15 : Bool;
         xSpare16 : Bool;
         xSpare17 : Bool;
         xSpare18 : Bool;
         xSpare19 : Bool;
         xSpare20 : Bool;
         xSpare21 : Bool;
         xSpare22 : Bool;
         xSpare23 : Bool;
         xSpare24 : Bool;
         xSpare25 : Bool;
         xSpare26 : Bool;
         xSpare27 : Bool;
         xSpare28 : Bool;
         xSpare29 : Bool;
         xSpare30 : Bool;
         xSpare31 : Bool;
         xSpare : Array[0..15] of Bool;
         iSpare0 : Int;
         iSpare1 : Int;
         iSpare2 : Int;
         iSpare3 : Int;
         iSpare4 : Int;
         iSpare5 : Int;
         iSpare6 : Int;
         iSpare7 : Int;
         iSpare8 : Int;
         iSpare9 : Int;
         iSpare10 : Int;
         iSpare11 : Int;
         iSpare12 : Int;
         iSpare13 : Int;
         iSpare14 : Int;
         iSpare15 : Int;
         iSpare16 : Int;
         dSpare0 : DInt;
         dSpare1 : DInt;
         dSpare2 : DInt;
         dSpare3 : DInt;
         dSpare4 : DInt;
         dSpare5 : DInt;
         dSpare6 : DInt;
         dSpare7 : DInt;
         dSpare8 : DInt;
         dSpare9 : DInt;
         dSpare10 : DInt;
         dSpare11 : DInt;
         dSpare12 : DInt;
         dSpare13 : DInt;
         dSpare14 : DInt;
         dSpare15 : DInt;
         rSpare0 : Real;
         rSpare1 : Real;
         rSpare2 : Real;
         rSpare3 : Real;
         rSpare4 : Real;
         rSpare5 : Real;
         rSpare6 : Real;
         rSpare7 : Real;
         rSpare8 : Real;
         tManCmd : Struct
            xSpare0 : Bool;
            xSpare1 : Bool;
            xSpare2 : Bool;
            xSpare3 : Bool;
            xSpare4 : Bool;
            xSpare5 : Bool;
            xSpare6 : Bool;
            xSpare7 : Bool;
            xSpare8 : Bool;
            xSpare9 : Bool;
            xSpare10 : Bool;
            xSpare11 : Bool;
            xSpare12 : Bool;
            xSpare13 : Bool;
            xSpare14 : Bool;
            xSpare15 : Bool;
            xSpare : Array[0..15] of Bool;
         END_STRUCT;
      END_STRUCT;
      tHMW : Struct   // HMI Write
         xSpare0 : Bool;
         xSpare1 : Bool;
         xSpare2 : Bool;
         xSpare3 : Bool;
         xSpare4 : Bool;
         xSpare5 : Bool;
         xSpare6 : Bool;
         xSpare7 : Bool;
         xSpare8 : Bool;
         xSpare9 : Bool;
         xSpare10 : Bool;
         xSpare11 : Bool;
         xSpare12 : Bool;
         xSpare13 : Bool;
         xSpare14 : Bool;
         xSpare15 : Bool;
         xSpare16 : Bool;
         xSpare17 : Bool;
         xSpare18 : Bool;
         xSpare19 : Bool;
         xSpare20 : Bool;
         xSpare21 : Bool;
         xSpare22 : Bool;
         xSpare23 : Bool;
         xSpare24 : Bool;
         xSpare25 : Bool;
         xSpare26 : Bool;
         xSpare27 : Bool;
         xSpare28 : Bool;
         xSpare29 : Bool;
         xSpare30 : Bool;
         xSpare31 : Bool;
         xSpare : Array[0..15] of Bool;
         iSpare0 : Int;
         iSpare1 : Int;
         iSpare2 : Int;
         iSpare3 : Int;
         iSpare4 : Int;
         iSpare5 : Int;
         iSpare6 : Int;
         iSpare7 : Int;
         iSpare8 : Int;
         iSpare9 : Int;
         iSpare10 : Int;
         iSpare11 : Int;
         iSpare12 : Int;
         iSpare13 : Int;
         iSpare14 : Int;
         iSpare15 : Int;
         iSpare16 : Int;
         dSpare0 : DInt;
         dSpare1 : DInt;
         dSpare2 : DInt;
         dSpare3 : DInt;
         dSpare4 : DInt;
         dSpare5 : DInt;
         dSpare6 : DInt;
         dSpare7 : DInt;
         dSpare8 : DInt;
         dSpare9 : DInt;
         dSpare10 : DInt;
         dSpare11 : DInt;
         dSpare12 : DInt;
         dSpare13 : DInt;
         dSpare14 : DInt;
         dSpare15 : DInt;
         dSpare16 : DInt;
         rSpare0 : Real;
         rSpare1 : Real;
         rSpare2 : Real;
         rSpare3 : Real;
         rSpare4 : Real;
         rSpare5 : Real;
         rSpare6 : Real;
         rSpare7 : Real;
         rSpare8 : Real;
         tManCmd : Struct
            xSpare0 : Bool;
            xSpare1 : Bool := false;
            xSpare2 : Bool;
            xSpare3 : Bool;
            xSpare4 : Bool;
            xSpare5 : Bool;
            xSpare6 : Bool;
            xSpare7 : Bool;
            xSpare8 : Bool;
            xSpare9 : Bool;
            xSpare10 : Bool;
            xSpare11 : Bool;
            xSpare12 : Bool;
            xSpare13 : Bool;
            xSpare14 : Bool;
            xSpare15 : Bool;
            xSpare16 : Bool;
            xSpare17 : Bool;
            xSpare18 : Bool;
            xSpare19 : Bool;
            xSpare20 : Bool;
            xSpare21 : Bool;
            xSpare22 : Bool;
            xSpare23 : Bool;
            xSpare24 : Bool;
            xSpare25 : Bool;
            xSpare26 : Bool;
            xSpare27 : Bool;
            xSpare28 : Bool;
            xSpare29 : Bool;
            xSpare30 : Bool;
            xSpare31 : Bool;
         END_STRUCT;
      END_STRUCT;
   END_VAR
BEGIN
END_DATA_BLOCK

DATA_BLOCK "DB_BPS_B_HMI"   // DB2111
{ S7_Optimized_Access := 'FALSE' }